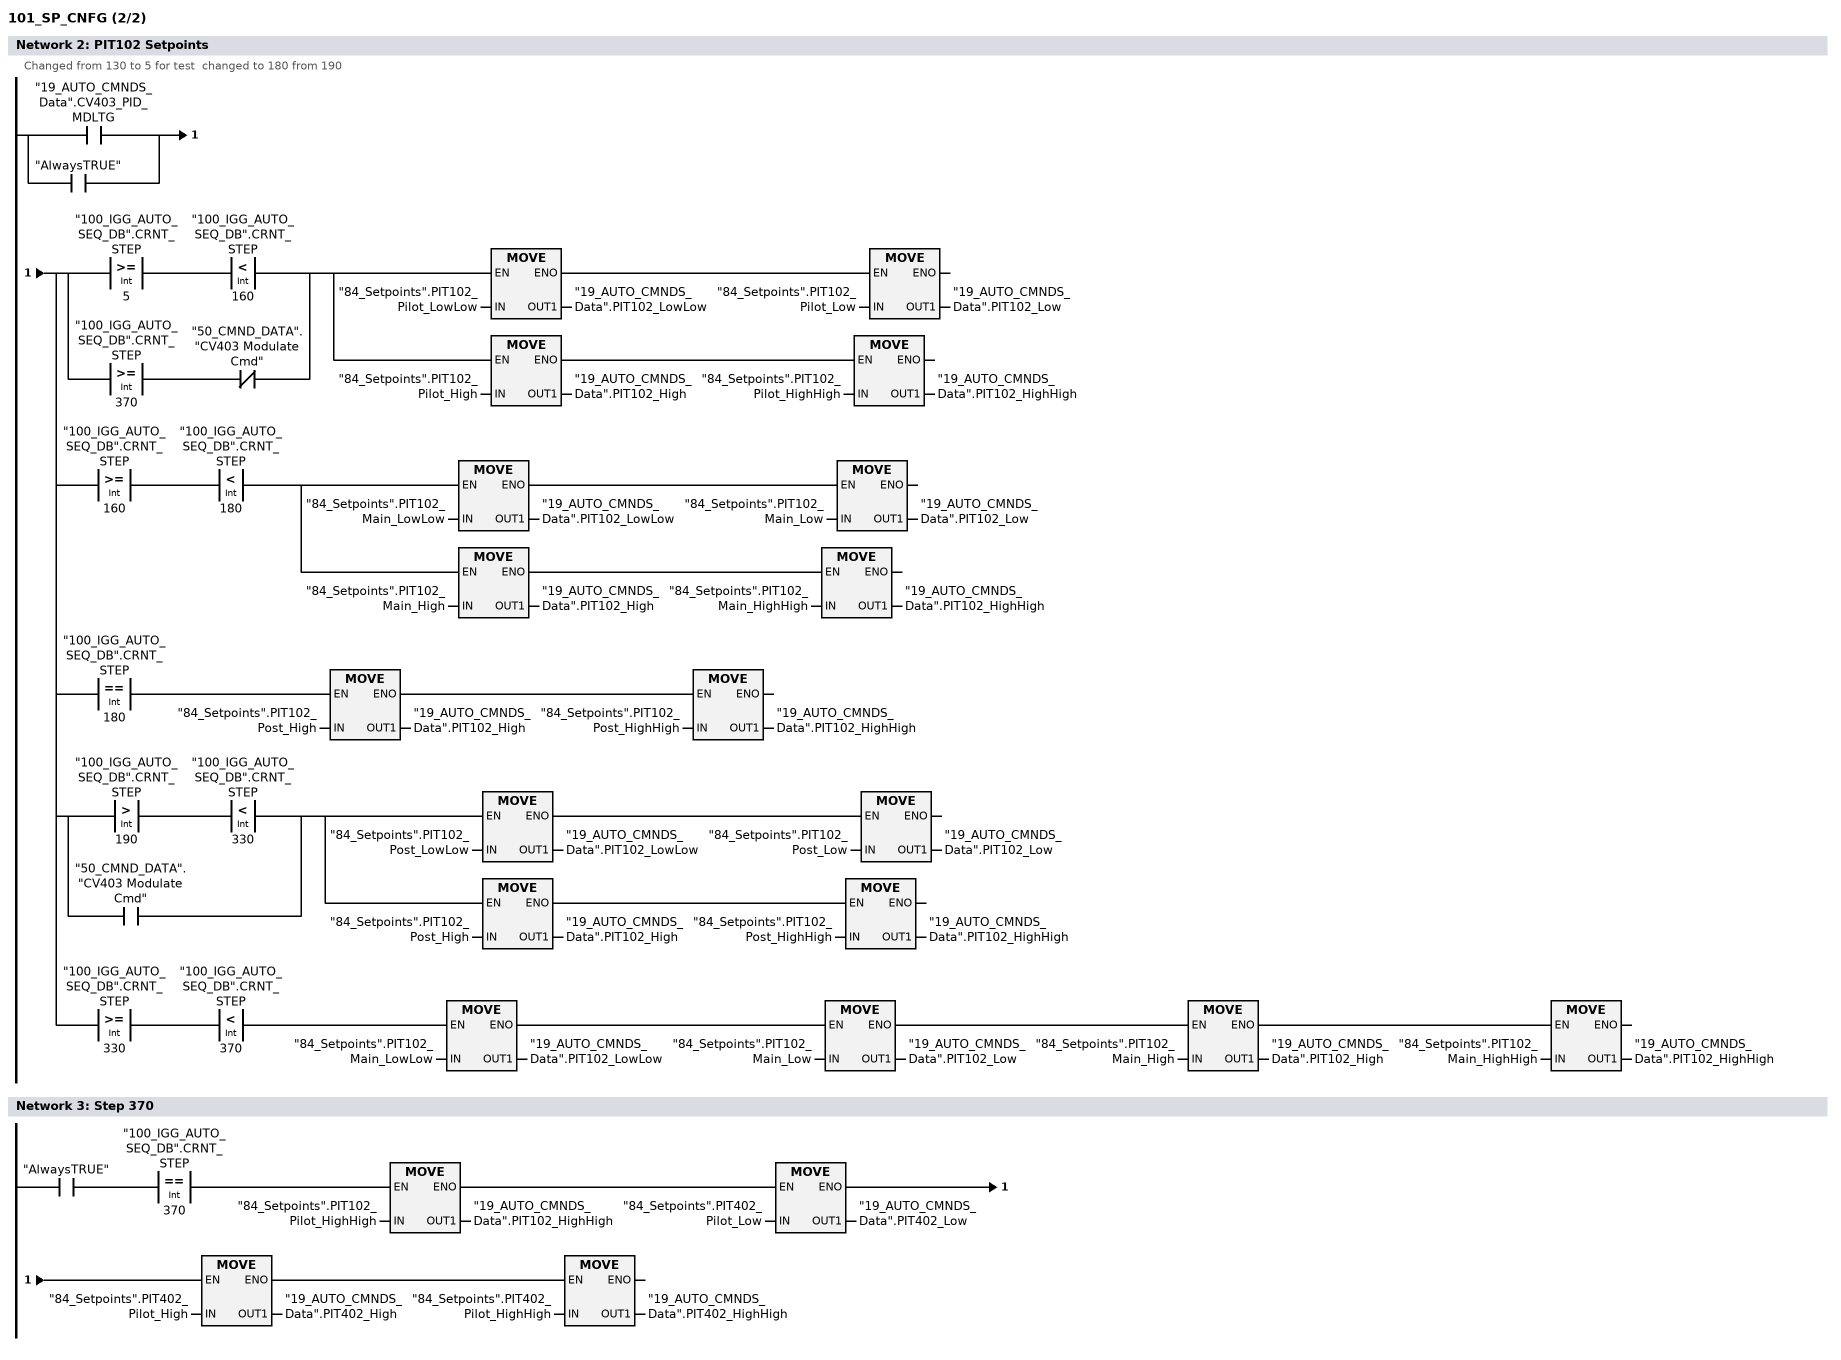
   RUNG wire#powerrail
      Contact( "19_AUTO_CMNDS_Data".CV403_PID_MDLTG )
      wire#w1
      { S7_Templates := "SrcType := Int" } GE_Contact(in1 := "100_IGG_AUTO_SEQ_DB".CRNT_STEP, in2 := 5)
      { S7_Templates := "SrcType := Int" } LT_Contact(in1 := "100_IGG_AUTO_SEQ_DB".CRNT_STEP, in2 := 160)
      wire#w2
      Move(in := "84_Setpoints".PIT102_Pilot_LowLow, out1 => "19_AUTO_CMNDS_Data".PIT102_LowLow)
      Move(in := "84_Setpoints".PIT102_Pilot_Low, out1 => "19_AUTO_CMNDS_Data".PIT102_Low)
   END_RUNG
   RUNG wire#powerrail
      Contact( "AlwaysTRUE" )
   END_RUNG wire#w1
   RUNG wire#w1
      { S7_Templates := "SrcType := Int" } GE_Contact(in1 := "100_IGG_AUTO_SEQ_DB".CRNT_STEP, in2 := 370)
      I_Contact( "50_CMND_DATA"."CV403 Modulate Cmd" )
   END_RUNG wire#w2
   RUNG wire#w2
      Move(in := "84_Setpoints".PIT102_Pilot_High, out1 => "19_AUTO_CMNDS_Data".PIT102_High)
      Move(in := "84_Setpoints".PIT102_Pilot_HighHigh, out1 => "19_AUTO_CMNDS_Data".PIT102_HighHigh)
   END_RUNG
   RUNG wire#w1
      { S7_Templates := "SrcType := Int" } GE_Contact(in1 := "100_IGG_AUTO_SEQ_DB".CRNT_STEP, in2 := 160)
      { S7_Templates := "SrcType := Int" } LT_Contact(in1 := "100_IGG_AUTO_SEQ_DB".CRNT_STEP, in2 := 180)
      wire#w3
      Move(in := "84_Setpoints".PIT102_Main_LowLow, out1 => "19_AUTO_CMNDS_Data".PIT102_LowLow)
      Move(in := "84_Setpoints".PIT102_Main_Low, out1 => "19_AUTO_CMNDS_Data".PIT102_Low)
   END_RUNG
   RUNG wire#w3
      Move(in := "84_Setpoints".PIT102_Main_High, out1 => "19_AUTO_CMNDS_Data".PIT102_High)
      Move(in := "84_Setpoints".PIT102_Main_HighHigh, out1 => "19_AUTO_CMNDS_Data".PIT102_HighHigh)
   END_RUNG
   RUNG wire#w1
      { S7_Templates := "SrcType := Int" } EQ_Contact(in1 := "100_IGG_AUTO_SEQ_DB".CRNT_STEP, in2 := 180)
      Move(in := "84_Setpoints".PIT102_Post_High, out1 => "19_AUTO_CMNDS_Data".PIT102_High)
      Move(in := "84_Setpoints".PIT102_Post_HighHigh, out1 => "19_AUTO_CMNDS_Data".PIT102_HighHigh)
   END_RUNG
   RUNG wire#w1
      { S7_Templates := "SrcType := Int" } GT_Contact(in1 := "100_IGG_AUTO_SEQ_DB".CRNT_STEP, in2 := 190)
      { S7_Templates := "SrcType := Int" } LT_Contact(in1 := "100_IGG_AUTO_SEQ_DB".CRNT_STEP, in2 := 330)
      wire#w4
      Move(in := "84_Setpoints".PIT102_Post_LowLow, out1 => "19_AUTO_CMNDS_Data".PIT102_LowLow)
      Move(in := "84_Setpoints".PIT102_Post_Low, out1 => "19_AUTO_CMNDS_Data".PIT102_Low)
   END_RUNG
   RUNG wire#w1
      Contact( "50_CMND_DATA"."CV403 Modulate Cmd" )
   END_RUNG wire#w4
   RUNG wire#w4
      Move(in := "84_Setpoints".PIT102_Post_High, out1 => "19_AUTO_CMNDS_Data".PIT102_High)
      Move(in := "84_Setpoints".PIT102_Post_HighHigh, out1 => "19_AUTO_CMNDS_Data".PIT102_HighHigh)
   END_RUNG
   RUNG wire#w1
      { S7_Templates := "SrcType := Int" } GE_Contact(in1 := "100_IGG_AUTO_SEQ_DB".CRNT_STEP, in2 := 330)
      { S7_Templates := "SrcType := Int" } LT_Contact(in1 := "100_IGG_AUTO_SEQ_DB".CRNT_STEP, in2 := 370)
      Move(in := "84_Setpoints".PIT102_Main_LowLow, out1 => "19_AUTO_CMNDS_Data".PIT102_LowLow)
      Move(in := "84_Setpoints".PIT102_Main_Low, out1 => "19_AUTO_CMNDS_Data".PIT102_Low)
      Move(in := "84_Setpoints".PIT102_Main_High, out1 => "19_AUTO_CMNDS_Data".PIT102_High)
      Move(in := "84_Setpoints".PIT102_Main_HighHigh, out1 => "19_AUTO_CMNDS_Data".PIT102_HighHigh)
   END_RUNG
   // the same network as SCL:
   #_w1 := "19_AUTO_CMNDS_Data".CV403_PID_MDLTG OR "AlwaysTRUE";
   IF #_w1 AND ((("100_IGG_AUTO_SEQ_DB".CRNT_STEP >= 5) AND ("100_IGG_AUTO_SEQ_DB".CRNT_STEP < 160)) OR (("100_IGG_AUTO_SEQ_DB".CRNT_STEP >= 370) AND NOT "50_CMND_DATA"."CV403 Modulate Cmd")) THEN
       "19_AUTO_CMNDS_Data".PIT102_LowLow := "84_Setpoints".PIT102_Pilot_LowLow;
       "19_AUTO_CMNDS_Data".PIT102_Low := "84_Setpoints".PIT102_Pilot_Low;
       "19_AUTO_CMNDS_Data".PIT102_High := "84_Setpoints".PIT102_Pilot_High;
       "19_AUTO_CMNDS_Data".PIT102_HighHigh := "84_Setpoints".PIT102_Pilot_HighHigh;
   END_IF;
   IF #_w1 AND ("100_IGG_AUTO_SEQ_DB".CRNT_STEP >= 160) AND ("100_IGG_AUTO_SEQ_DB".CRNT_STEP < 180) THEN
       "19_AUTO_CMNDS_Data".PIT102_LowLow := "84_Setpoints".PIT102_Main_LowLow;
       "19_AUTO_CMNDS_Data".PIT102_Low := "84_Setpoints".PIT102_Main_Low;
       "19_AUTO_CMNDS_Data".PIT102_High := "84_Setpoints".PIT102_Main_High;
       "19_AUTO_CMNDS_Data".PIT102_HighHigh := "84_Setpoints".PIT102_Main_HighHigh;
   END_IF;
   IF #_w1 AND ("100_IGG_AUTO_SEQ_DB".CRNT_STEP = 180) THEN
       "19_AUTO_CMNDS_Data".PIT102_High := "84_Setpoints".PIT102_Post_High;
       "19_AUTO_CMNDS_Data".PIT102_HighHigh := "84_Setpoints".PIT102_Post_HighHigh;
   END_IF;
   IF #_w1 AND ((("100_IGG_AUTO_SEQ_DB".CRNT_STEP > 190) AND ("100_IGG_AUTO_SEQ_DB".CRNT_STEP < 330)) OR "50_CMND_DATA"."CV403 Modulate Cmd") THEN
       "19_AUTO_CMNDS_Data".PIT102_LowLow := "84_Setpoints".PIT102_Post_LowLow;
       "19_AUTO_CMNDS_Data".PIT102_Low := "84_Setpoints".PIT102_Post_Low;
       "19_AUTO_CMNDS_Data".PIT102_High := "84_Setpoints".PIT102_Post_High;
       "19_AUTO_CMNDS_Data".PIT102_HighHigh := "84_Setpoints".PIT102_Post_HighHigh;
   END_IF;
   IF #_w1 AND ("100_IGG_AUTO_SEQ_DB".CRNT_STEP >= 330) AND ("100_IGG_AUTO_SEQ_DB".CRNT_STEP < 370) THEN
       "19_AUTO_CMNDS_Data".PIT102_LowLow := "84_Setpoints".PIT102_Main_LowLow;
       "19_AUTO_CMNDS_Data".PIT102_Low := "84_Setpoints".PIT102_Main_Low;
       "19_AUTO_CMNDS_Data".PIT102_High := "84_Setpoints".PIT102_Main_High;
       "19_AUTO_CMNDS_Data".PIT102_HighHigh := "84_Setpoints".PIT102_Main_HighHigh;
   END_IF;
END_REGION

REGION Network 3: Step 370
   RUNG wire#powerrail
      Contact( "AlwaysTRUE" )
      { S7_Templates := "SrcType := Int" } EQ_Contact(in1 := "100_IGG_AUTO_SEQ_DB".CRNT_STEP, in2 := 370)
      Move(in := "84_Setpoints".PIT102_Pilot_HighHigh, out1 => "19_AUTO_CMNDS_Data".PIT102_HighHigh)
      Move(in := "84_Setpoints".PIT402_Pilot_Low, out1 => "19_AUTO_CMNDS_Data".PIT402_Low)
      Move(in := "84_Setpoints".PIT402_Pilot_High, out1 => "19_AUTO_CMNDS_Data".PIT402_High)
      Move(in := "84_Setpoints".PIT402_Pilot_HighHigh, out1 => "19_AUTO_CMNDS_Data".PIT402_HighHigh)
   END_RUNG
   // the same network as SCL:
   IF "AlwaysTRUE" AND ("100_IGG_AUTO_SEQ_DB".CRNT_STEP = 370) THEN
       "19_AUTO_CMNDS_Data".PIT102_HighHigh := "84_Setpoints".PIT102_Pilot_HighHigh;
       "19_AUTO_CMNDS_Data".PIT402_Low := "84_Setpoints".PIT402_Pilot_Low;
       "19_AUTO_CMNDS_Data".PIT402_High := "84_Setpoints".PIT402_Pilot_High;
       "19_AUTO_CMNDS_Data".PIT402_HighHigh := "84_Setpoints".PIT402_Pilot_HighHigh;
   END_IF;
END_REGION
END_FUNCTION

// folder: 120 - 139 FAT Functions

FUNCTION "120_FAT_FCS" : Void   // FC120, LAD
TITLE = FAT Functions
{ S7_Optimized_Access := 'TRUE' }
AUTHOR : JRS
VERSION : 0.1
// For specific functions related to the factory test equipment & setup
   VAR_TEMP   // added for the SCL form of the ladder/FBD networks
      _w1 : Bool;
   END_VAR
BEGIN

REGION Network 1: Into FAT Mode
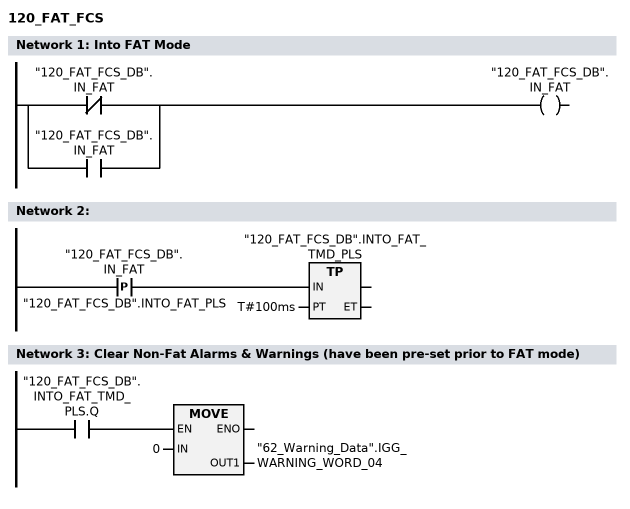
   RUNG wire#powerrail
      I_Contact( "120_FAT_FCS_DB".IN_FAT )
      wire#w1
      Coil( "120_FAT_FCS_DB".IN_FAT )
   END_RUNG
   RUNG wire#powerrail
      Contact( "120_FAT_FCS_DB".IN_FAT )
   END_RUNG wire#w1
   // the same network as SCL:
   "120_FAT_FCS_DB".IN_FAT := NOT "120_FAT_FCS_DB".IN_FAT OR "120_FAT_FCS_DB".IN_FAT;
END_REGION

REGION Network 2
   #_w1 := "120_FAT_FCS_DB".IN_FAT AND NOT "120_FAT_FCS_DB".INTO_FAT_PLS;   // rising edge of "120_FAT_FCS_DB".IN_FAT
   "120_FAT_FCS_DB".INTO_FAT_PLS := "120_FAT_FCS_DB".IN_FAT;
   "120_FAT_FCS_DB".INTO_FAT_TMD_PLS.TP(IN := #_w1, PT := T#100ms);
END_REGION

REGION Network 3: Clear Non-Fat Alarms & Warnings (have been pre-set prior to FAT mode)
   RUNG wire#powerrail
      Contact( "120_FAT_FCS_DB".INTO_FAT_TMD_PLS.Q )
      Move(in := 0, out1 => "62_Warning_Data".IGG_WARNING_WORD_04)
   END_RUNG
   // the same network as SCL:
   IF "120_FAT_FCS_DB".INTO_FAT_TMD_PLS.Q THEN "62_Warning_Data".IGG_WARNING_WORD_04 := 0; END_IF;
END_REGION
END_FUNCTION

// folder: 300 - 499 Counters and Timer DBs

FUNCTION "300_AUT_SUQ_TIMERS" : Void   // FC300, LAD
TITLE = Automatic Sequence Timers
{ S7_Optimized_Access := 'TRUE' }
AUTHOR : JRS
VERSION : 0.1
// For specific sequence timers not covered by step FB timers
BEGIN

REGION Network 1: Pre BC Start Command Delay
   // Get time value from HMI data
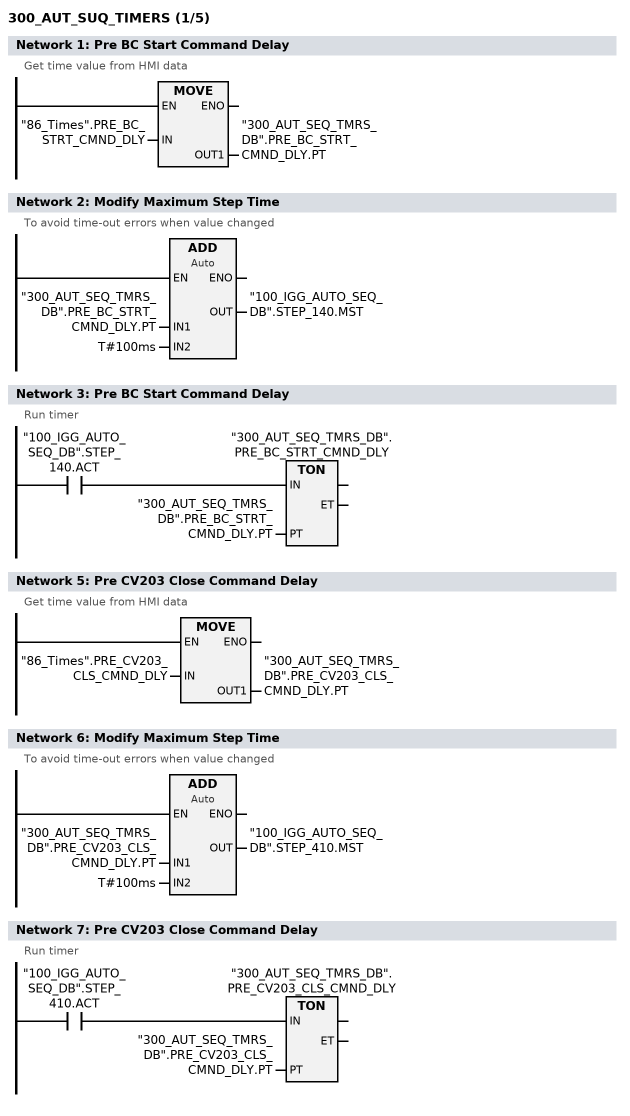
   RUNG wire#powerrail
      Move(in := "86_Times".PRE_BC_STRT_CMND_DLY, out1 => "300_AUT_SEQ_TMRS_DB".PRE_BC_STRT_CMND_DLY.PT)
   END_RUNG
   // the same network as SCL:
   "300_AUT_SEQ_TMRS_DB".PRE_BC_STRT_CMND_DLY.PT := "86_Times".PRE_BC_STRT_CMND_DLY;
END_REGION

REGION Network 2: Modify Maximum Step Time
   // To avoid time-out errors when value changed
   RUNG wire#powerrail
      Add(in1 := "300_AUT_SEQ_TMRS_DB".PRE_BC_STRT_CMND_DLY.PT, in2 := T#100ms, out => "100_IGG_AUTO_SEQ_DB".STEP_140.MST)
   END_RUNG
   // the same network as SCL:
   "100_IGG_AUTO_SEQ_DB".STEP_140.MST := "300_AUT_SEQ_TMRS_DB".PRE_BC_STRT_CMND_DLY.PT + T#100ms;
END_REGION

REGION Network 3: Pre BC Start Command Delay
   // Run timer
   "300_AUT_SEQ_TMRS_DB".PRE_BC_STRT_CMND_DLY.TON(IN := "100_IGG_AUTO_SEQ_DB".STEP_140.ACT,
                           PT := "300_AUT_SEQ_TMRS_DB".PRE_BC_STRT_CMND_DLY.PT);
END_REGION

REGION Network 5: Pre CV203 Close Command Delay
   // Get time value from HMI data
   RUNG wire#powerrail
      Move(in := "86_Times".PRE_CV203_CLS_CMND_DLY, out1 => "300_AUT_SEQ_TMRS_DB".PRE_CV203_CLS_CMND_DLY.PT)
   END_RUNG
   // the same network as SCL:
   "300_AUT_SEQ_TMRS_DB".PRE_CV203_CLS_CMND_DLY.PT := "86_Times".PRE_CV203_CLS_CMND_DLY;
END_REGION

REGION Network 6: Modify Maximum Step Time
   // To avoid time-out errors when value changed
   RUNG wire#powerrail
      Add(in1 := "300_AUT_SEQ_TMRS_DB".PRE_CV203_CLS_CMND_DLY.PT, in2 := T#100ms, out => "100_IGG_AUTO_SEQ_DB".STEP_410.MST)
   END_RUNG
   // the same network as SCL:
   "100_IGG_AUTO_SEQ_DB".STEP_410.MST := "300_AUT_SEQ_TMRS_DB".PRE_CV203_CLS_CMND_DLY.PT + T#100ms;
END_REGION

REGION Network 7: Pre CV203 Close Command Delay
   // Run timer
   "300_AUT_SEQ_TMRS_DB".PRE_CV203_CLS_CMND_DLY.TON(IN := "100_IGG_AUTO_SEQ_DB".STEP_410.ACT,
                           PT := "300_AUT_SEQ_TMRS_DB".PRE_CV203_CLS_CMND_DLY.PT);
END_REGION

REGION Network 9: Post P301 Stop Delay
   // Get time value from HMI data
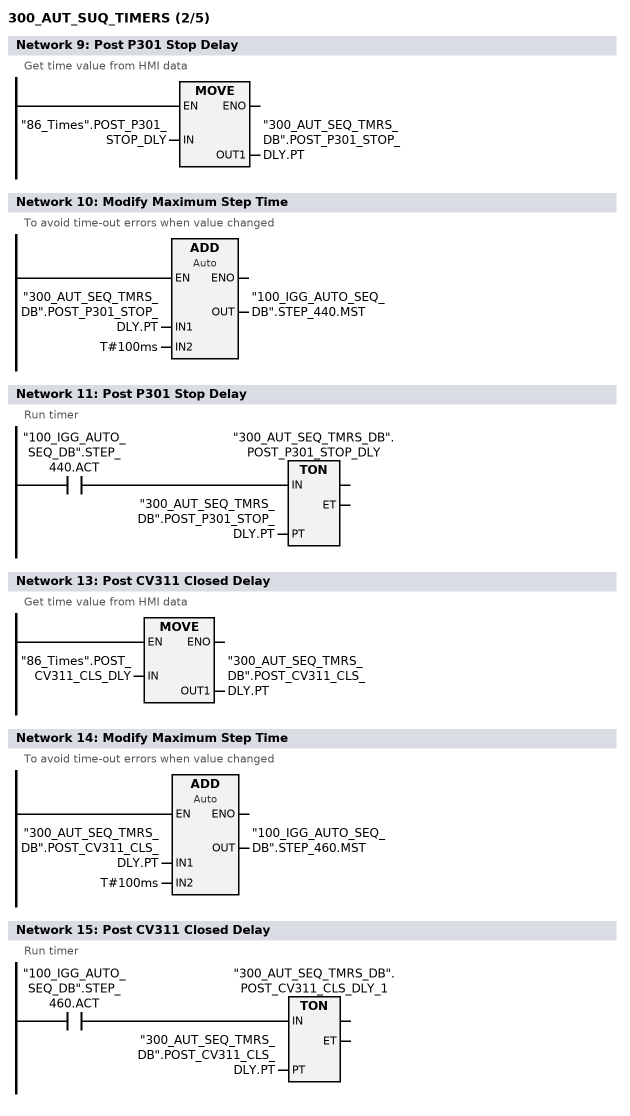
   RUNG wire#powerrail
      Move(in := "86_Times".POST_P301_STOP_DLY, out1 => "300_AUT_SEQ_TMRS_DB".POST_P301_STOP_DLY.PT)
   END_RUNG
   // the same network as SCL:
   "300_AUT_SEQ_TMRS_DB".POST_P301_STOP_DLY.PT := "86_Times".POST_P301_STOP_DLY;
END_REGION

REGION Network 10: Modify Maximum Step Time
   // To avoid time-out errors when value changed
   RUNG wire#powerrail
      Add(in1 := "300_AUT_SEQ_TMRS_DB".POST_P301_STOP_DLY.PT, in2 := T#100ms, out => "100_IGG_AUTO_SEQ_DB".STEP_440.MST)
   END_RUNG
   // the same network as SCL:
   "100_IGG_AUTO_SEQ_DB".STEP_440.MST := "300_AUT_SEQ_TMRS_DB".POST_P301_STOP_DLY.PT + T#100ms;
END_REGION

REGION Network 11: Post P301 Stop Delay
   // Run timer
   "300_AUT_SEQ_TMRS_DB".POST_P301_STOP_DLY.TON(IN := "100_IGG_AUTO_SEQ_DB".STEP_440.ACT,
                           PT := "300_AUT_SEQ_TMRS_DB".POST_P301_STOP_DLY.PT);
END_REGION

REGION Network 13: Post CV311 Closed Delay
   // Get time value from HMI data
   RUNG wire#powerrail
      Move(in := "86_Times".POST_CV311_CLS_DLY, out1 => "300_AUT_SEQ_TMRS_DB".POST_CV311_CLS_DLY.PT)
   END_RUNG
   // the same network as SCL:
   "300_AUT_SEQ_TMRS_DB".POST_CV311_CLS_DLY.PT := "86_Times".POST_CV311_CLS_DLY;
END_REGION

REGION Network 14: Modify Maximum Step Time
   // To avoid time-out errors when value changed
   RUNG wire#powerrail
      Add(in1 := "300_AUT_SEQ_TMRS_DB".POST_CV311_CLS_DLY.PT, in2 := T#100ms, out => "100_IGG_AUTO_SEQ_DB".STEP_460.MST)
   END_RUNG
   // the same network as SCL:
   "100_IGG_AUTO_SEQ_DB".STEP_460.MST := "300_AUT_SEQ_TMRS_DB".POST_CV311_CLS_DLY.PT + T#100ms;
END_REGION

REGION Network 15: Post CV311 Closed Delay
   // Run timer
   "300_AUT_SEQ_TMRS_DB".POST_CV311_CLS_DLY_1.TON(IN := "100_IGG_AUTO_SEQ_DB".STEP_460.ACT,
                           PT := "300_AUT_SEQ_TMRS_DB".POST_CV311_CLS_DLY.PT);
END_REGION

REGION Network 17: Post CV321 Opened Delay
   // Get time value from HMI data
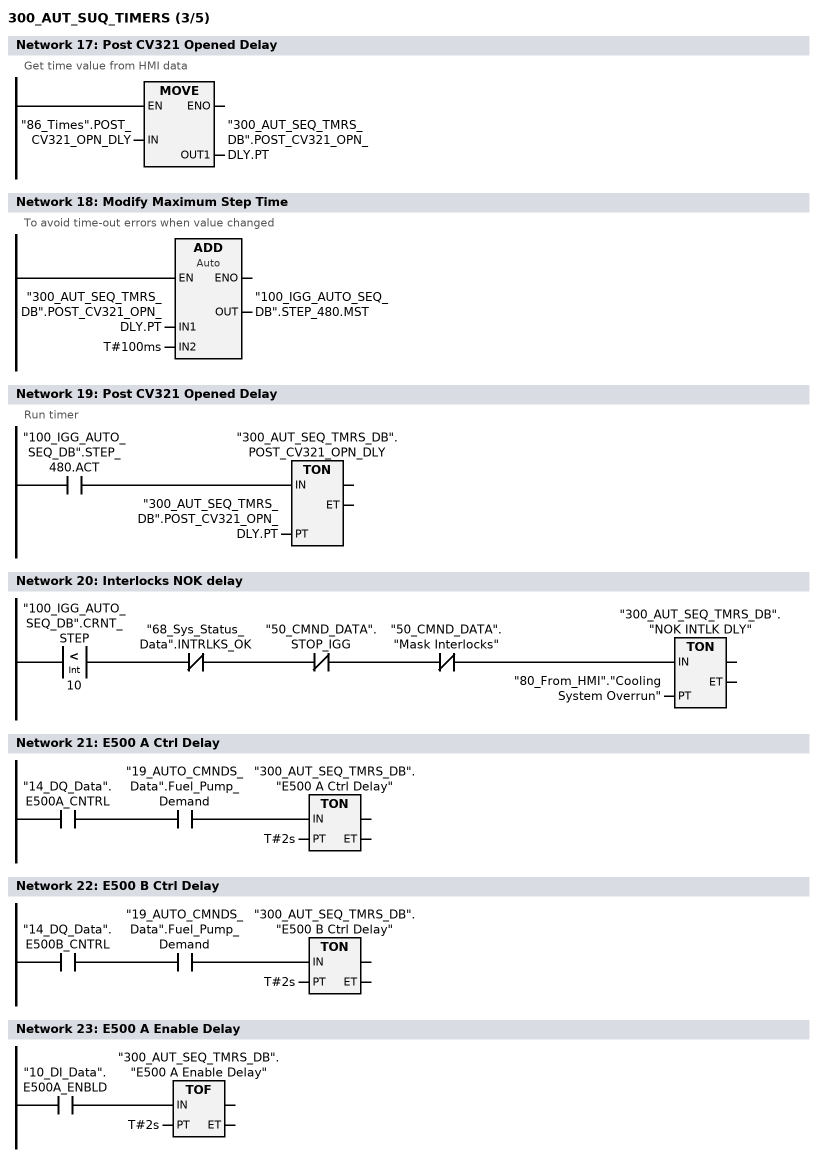
   RUNG wire#powerrail
      Move(in := "86_Times".POST_CV321_OPN_DLY, out1 => "300_AUT_SEQ_TMRS_DB".POST_CV321_OPN_DLY.PT)
   END_RUNG
   // the same network as SCL:
   "300_AUT_SEQ_TMRS_DB".POST_CV321_OPN_DLY.PT := "86_Times".POST_CV321_OPN_DLY;
END_REGION

REGION Network 18: Modify Maximum Step Time
   // To avoid time-out errors when value changed
   RUNG wire#powerrail
      Add(in1 := "300_AUT_SEQ_TMRS_DB".POST_CV321_OPN_DLY.PT, in2 := T#100ms, out => "100_IGG_AUTO_SEQ_DB".STEP_480.MST)
   END_RUNG
   // the same network as SCL:
   "100_IGG_AUTO_SEQ_DB".STEP_480.MST := "300_AUT_SEQ_TMRS_DB".POST_CV321_OPN_DLY.PT + T#100ms;
END_REGION

REGION Network 19: Post CV321 Opened Delay
   // Run timer
   "300_AUT_SEQ_TMRS_DB".POST_CV321_OPN_DLY.TON(IN := "100_IGG_AUTO_SEQ_DB".STEP_480.ACT,
                           PT := "300_AUT_SEQ_TMRS_DB".POST_CV321_OPN_DLY.PT);
END_REGION

REGION Network 20: Interlocks NOK delay
   "300_AUT_SEQ_TMRS_DB"."NOK INTLK DLY".TON(IN := ("100_IGG_AUTO_SEQ_DB".CRNT_STEP < 10) AND NOT "68_Sys_Status_Data".INTRLKS_OK AND NOT "50_CMND_DATA".STOP_IGG AND NOT "50_CMND_DATA"."Mask Interlocks",
                           PT := "80_From_HMI"."Cooling System Overrun");
END_REGION

REGION Network 21: E500 A Ctrl Delay
   "300_AUT_SEQ_TMRS_DB"."E500 A Ctrl Delay".TON(IN := "14_DQ_Data".E500A_CNTRL AND "19_AUTO_CMNDS_Data".Fuel_Pump_Demand,
                           PT := T#2s);
END_REGION

REGION Network 22: E500 B Ctrl Delay
   "300_AUT_SEQ_TMRS_DB"."E500 B Ctrl Delay".TON(IN := "14_DQ_Data".E500B_CNTRL AND "19_AUTO_CMNDS_Data".Fuel_Pump_Demand,
                           PT := T#2s);
END_REGION

REGION Network 23: E500 A Enable Delay
   "300_AUT_SEQ_TMRS_DB"."E500 A Enable Delay".TOF(IN := "10_DI_Data".E500A_ENBLD, PT := T#2s);
END_REGION

REGION Network 24: E500 B Enable Delay
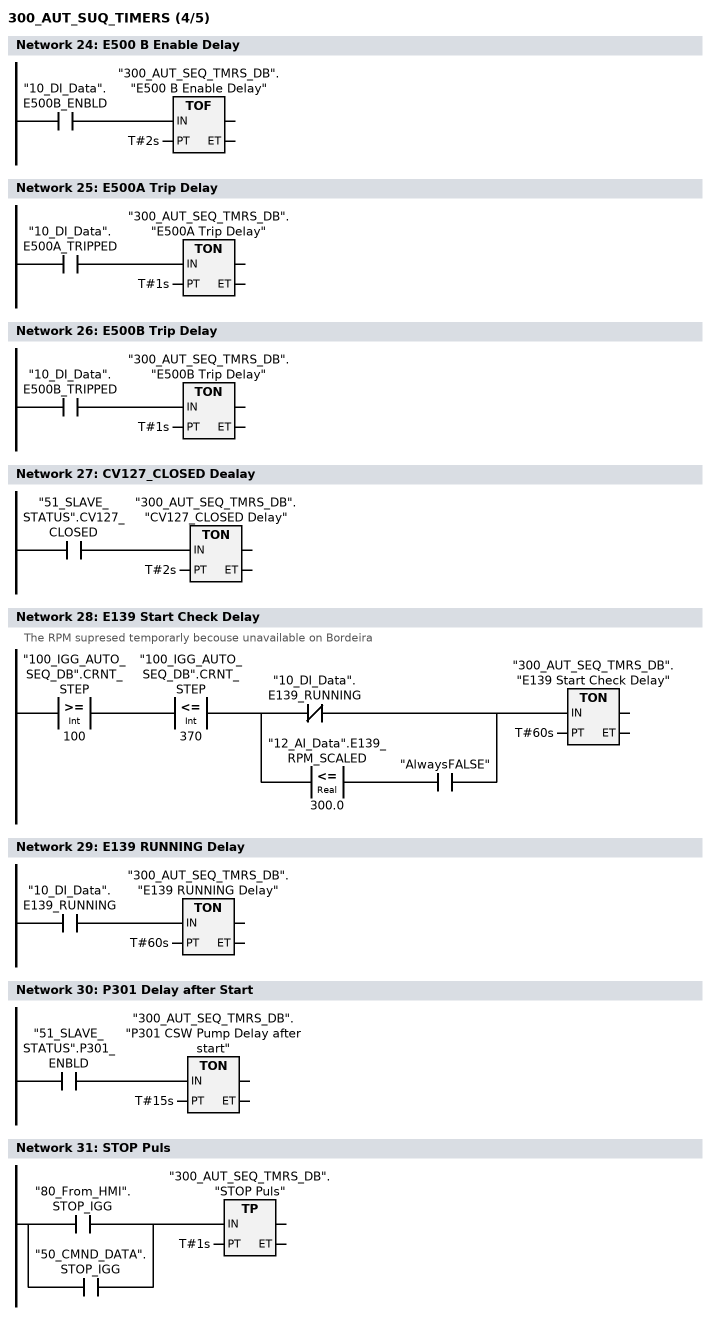
   "300_AUT_SEQ_TMRS_DB"."E500 B Enable Delay".TOF(IN := "10_DI_Data".E500B_ENBLD, PT := T#2s);
END_REGION

REGION Network 25: E500A Trip Delay
   "300_AUT_SEQ_TMRS_DB"."E500A Trip Delay".TON(IN := "10_DI_Data".E500A_TRIPPED, PT := T#1s);
END_REGION

REGION Network 26: E500B Trip Delay
   "300_AUT_SEQ_TMRS_DB"."E500B Trip Delay".TON(IN := "10_DI_Data".E500B_TRIPPED, PT := T#1s);
END_REGION

REGION Network 27: CV127_CLOSED Dealay
   "300_AUT_SEQ_TMRS_DB"."CV127_CLOSED Delay".TON(IN := "51_SLAVE_STATUS".CV127_CLOSED, PT := T#2s);
END_REGION

REGION Network 28: E139 Start Check Delay
   // The RPM supresed temporarly becouse unavailable on Bordeira
   "300_AUT_SEQ_TMRS_DB"."E139 Start Check Delay".TON(IN := ("100_IGG_AUTO_SEQ_DB".CRNT_STEP >= 100) AND ("100_IGG_AUTO_SEQ_DB".CRNT_STEP <= 370) AND (NOT "10_DI_Data".E139_RUNNING OR (("12_AI_Data".E139_RPM_SCALED <= 300.0) AND "AlwaysFALSE")),
                           PT := T#60s);
END_REGION

REGION Network 29: E139 RUNNING Delay
   "300_AUT_SEQ_TMRS_DB"."E139 RUNNING Delay".TON(IN := "10_DI_Data".E139_RUNNING, PT := T#60s);
END_REGION

REGION Network 30: P301 Delay after Start
   "300_AUT_SEQ_TMRS_DB"."P301 CSW Pump Delay after start".TON(IN := "51_SLAVE_STATUS".P301_ENBLD, PT := T#15s);
END_REGION

REGION Network 31: STOP Puls
   "300_AUT_SEQ_TMRS_DB"."STOP Puls".TP(IN := "80_From_HMI".STOP_IGG OR "50_CMND_DATA".STOP_IGG, PT := T#1s);
END_REGION

REGION Network 32: E-Stop Loop
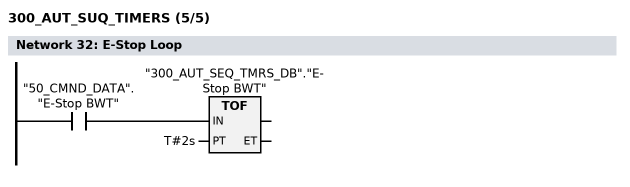
   "300_AUT_SEQ_TMRS_DB"."E-Stop BWT".TOF(IN := "50_CMND_DATA"."E-Stop BWT", PT := T#2s);
END_REGION
END_FUNCTION

// folder: 50 - 59 Communication

FUNCTION "51_GET_SLAVE_DATA" : Void   // FC51, LAD
TITLE = Get Slave Status Data
{ S7_Optimized_Access := 'TRUE' }
AUTHOR : JRS
VERSION : 0.1
// Code for getting status data from the slave PLC
BEGIN

REGION Network 1: Get Slave Status Data
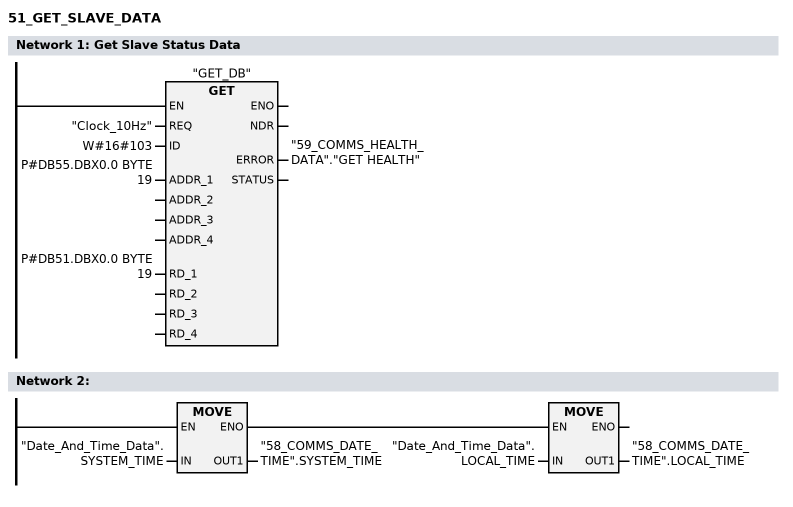
   "GET_DB"(REQ := "Clock_10Hz",   // GET
            ID := W#16#103,
            ADDR_1 := P#DB55.DBX0.0 BYTE 19,
            RD_1 := P#DB51.DBX0.0 BYTE 19,
            ERROR => "59_COMMS_HEALTH_DATA"."GET HEALTH");
END_REGION

REGION Network 2
   RUNG wire#powerrail
      Move(in := "Date_And_Time_Data".SYSTEM_TIME, out1 => "58_COMMS_DATE_TIME".SYSTEM_TIME)
      Move(in := "Date_And_Time_Data".LOCAL_TIME, out1 => "58_COMMS_DATE_TIME".LOCAL_TIME)
   END_RUNG
   // the same network as SCL:
   "58_COMMS_DATE_TIME".SYSTEM_TIME := "Date_And_Time_Data".SYSTEM_TIME;
   "58_COMMS_DATE_TIME".LOCAL_TIME := "Date_And_Time_Data".LOCAL_TIME;
END_REGION
END_FUNCTION

FUNCTION "56_PUT_SLAVE_DATA" : Void   // FC56, LAD
TITLE = Put Slave Comands Data
{ S7_Optimized_Access := 'TRUE' }
AUTHOR : JRS
VERSION : 0.1
// Code for sending commands to the slave PLC
   VAR_TEMP
      RACK_2_done : Bool;
      RACK_2_error : Bool;
      RACK_2_status : Word;
      RACK_3_done : Bool;
      RACK_3_error : Bool;
      RACK_3_status : Word;
   END_VAR
BEGIN

REGION Network 1: PUT Slave Commands
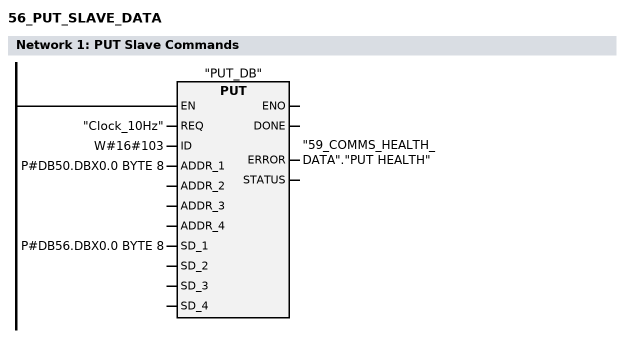
   "PUT_DB"(REQ := "Clock_10Hz",   // PUT
            ID := W#16#103,
            ADDR_1 := P#DB50.DBX0.0 BYTE 8,
            SD_1 := P#DB56.DBX0.0 BYTE 8,
            ERROR => "59_COMMS_HEALTH_DATA"."PUT HEALTH");
END_REGION
END_FUNCTION

FUNCTION "59_COMMS_HEALTH" : Void   // FC59, LAD
TITLE = Communications Heart Beats
{ S7_Optimized_Access := 'TRUE' }
AUTHOR : JRS
VERSION : 0.1
// Code for communications health determination
   VAR_TEMP   // added for the SCL form of the ladder/FBD networks
      _w1 : Bool;
      _w2 : Bool;
   END_VAR
BEGIN

REGION Network 1: Local Heart Beat
   // Flip flop for status to other PLC's
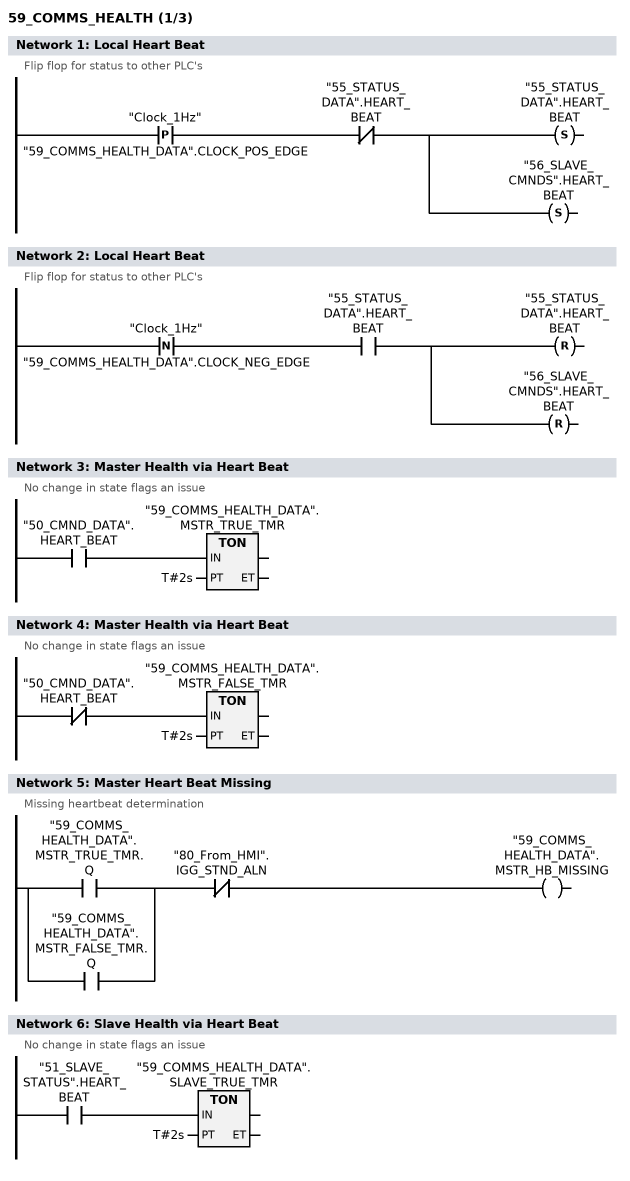
   RUNG wire#powerrail
      P_Contact(operand := "Clock_1Hz", bit := "59_COMMS_HEALTH_DATA".CLOCK_POS_EDGE)
      I_Contact( "55_STATUS_DATA".HEART_BEAT )
      wire#w1
      S_Coil( "55_STATUS_DATA".HEART_BEAT )
   END_RUNG
   RUNG wire#w1
      S_Coil( "56_SLAVE_CMNDS".HEART_BEAT )
   END_RUNG
   // the same network as SCL:
   #_w1 := "Clock_1Hz" AND NOT "59_COMMS_HEALTH_DATA".CLOCK_POS_EDGE;   // rising edge of "Clock_1Hz"
   "59_COMMS_HEALTH_DATA".CLOCK_POS_EDGE := "Clock_1Hz";
   #_w2 := #_w1 AND NOT "55_STATUS_DATA".HEART_BEAT;
   IF #_w2 THEN
       "55_STATUS_DATA".HEART_BEAT := TRUE;
       "56_SLAVE_CMNDS".HEART_BEAT := TRUE;
   END_IF;
END_REGION

REGION Network 2: Local Heart Beat
   // Flip flop for status to other PLC's
   RUNG wire#powerrail
      N_Contact(operand := "Clock_1Hz", bit := "59_COMMS_HEALTH_DATA".CLOCK_NEG_EDGE)
      Contact( "55_STATUS_DATA".HEART_BEAT )
      wire#w1
      R_Coil( "55_STATUS_DATA".HEART_BEAT )
   END_RUNG
   RUNG wire#w1
      R_Coil( "56_SLAVE_CMNDS".HEART_BEAT )
   END_RUNG
   // the same network as SCL:
   #_w1 := NOT "Clock_1Hz" AND "59_COMMS_HEALTH_DATA".CLOCK_NEG_EDGE;   // falling edge of "Clock_1Hz"
   "59_COMMS_HEALTH_DATA".CLOCK_NEG_EDGE := "Clock_1Hz";
   #_w2 := #_w1 AND "55_STATUS_DATA".HEART_BEAT;
   IF #_w2 THEN
       "55_STATUS_DATA".HEART_BEAT := FALSE;
       "56_SLAVE_CMNDS".HEART_BEAT := FALSE;
   END_IF;
END_REGION

REGION Network 3: Master Health via Heart Beat
   // No change in state flags an issue
   "59_COMMS_HEALTH_DATA".MSTR_TRUE_TMR.TON(IN := "50_CMND_DATA".HEART_BEAT, PT := T#2s);
END_REGION

REGION Network 4: Master Health via Heart Beat
   // No change in state flags an issue
   "59_COMMS_HEALTH_DATA".MSTR_FALSE_TMR.TON(IN := NOT "50_CMND_DATA".HEART_BEAT, PT := T#2s);
END_REGION

REGION Network 5: Master Heart Beat Missing
   // Missing heartbeat determination
   RUNG wire#powerrail
      Contact( "59_COMMS_HEALTH_DATA".MSTR_TRUE_TMR.Q )
      wire#w1
      I_Contact( "80_From_HMI".IGG_STND_ALN )
      Coil( "59_COMMS_HEALTH_DATA".MSTR_HB_MISSING )
   END_RUNG
   RUNG wire#powerrail
      Contact( "59_COMMS_HEALTH_DATA".MSTR_FALSE_TMR.Q )
   END_RUNG wire#w1
   // the same network as SCL:
   "59_COMMS_HEALTH_DATA".MSTR_HB_MISSING := ("59_COMMS_HEALTH_DATA".MSTR_TRUE_TMR.Q OR "59_COMMS_HEALTH_DATA".MSTR_FALSE_TMR.Q) AND NOT "80_From_HMI".IGG_STND_ALN;
END_REGION

REGION Network 6: Slave Health via Heart Beat
   // No change in state flags an issue
   "59_COMMS_HEALTH_DATA".SLAVE_TRUE_TMR.TON(IN := "51_SLAVE_STATUS".HEART_BEAT, PT := T#2s);
END_REGION

REGION Network 7: Slave Health via Heart Beat
   // No change in state flags an issue
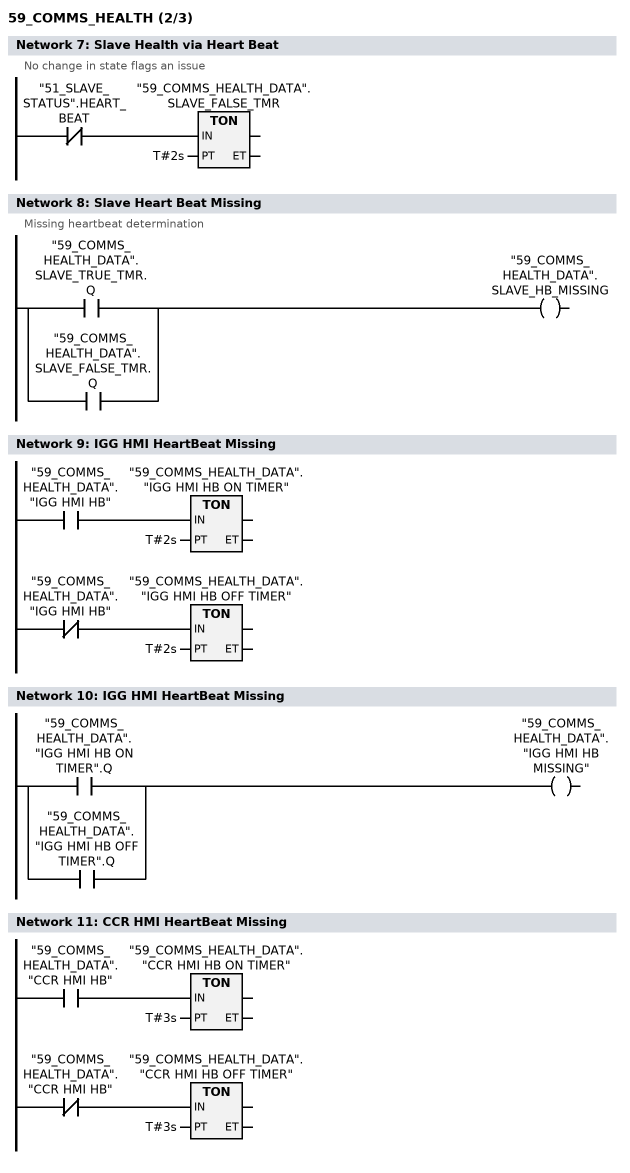
   "59_COMMS_HEALTH_DATA".SLAVE_FALSE_TMR.TON(IN := NOT "51_SLAVE_STATUS".HEART_BEAT, PT := T#2s);
END_REGION

REGION Network 8: Slave Heart Beat Missing
   // Missing heartbeat determination
   RUNG wire#powerrail
      Contact( "59_COMMS_HEALTH_DATA".SLAVE_TRUE_TMR.Q )
      wire#w1
      Coil( "59_COMMS_HEALTH_DATA".SLAVE_HB_MISSING )
   END_RUNG
   RUNG wire#powerrail
      Contact( "59_COMMS_HEALTH_DATA".SLAVE_FALSE_TMR.Q )
   END_RUNG wire#w1
   // the same network as SCL:
   "59_COMMS_HEALTH_DATA".SLAVE_HB_MISSING := "59_COMMS_HEALTH_DATA".SLAVE_TRUE_TMR.Q OR "59_COMMS_HEALTH_DATA".SLAVE_FALSE_TMR.Q;
END_REGION

REGION Network 9: IGG HMI HeartBeat Missing
   "59_COMMS_HEALTH_DATA"."IGG HMI HB ON TIMER".TON(IN := "59_COMMS_HEALTH_DATA"."IGG HMI HB", PT := T#2s);
   "59_COMMS_HEALTH_DATA"."IGG HMI HB OFF TIMER".TON(IN := NOT "59_COMMS_HEALTH_DATA"."IGG HMI HB", PT := T#2s);
END_REGION

REGION Network 10: IGG HMI HeartBeat Missing
   RUNG wire#powerrail
      Contact( "59_COMMS_HEALTH_DATA"."IGG HMI HB ON TIMER".Q )
      wire#w1
      Coil( "59_COMMS_HEALTH_DATA"."IGG HMI HB MISSING" )
   END_RUNG
   RUNG wire#powerrail
      Contact( "59_COMMS_HEALTH_DATA"."IGG HMI HB OFF TIMER".Q )
   END_RUNG wire#w1
   // the same network as SCL:
   "59_COMMS_HEALTH_DATA"."IGG HMI HB MISSING" := "59_COMMS_HEALTH_DATA"."IGG HMI HB ON TIMER".Q OR "59_COMMS_HEALTH_DATA"."IGG HMI HB OFF TIMER".Q;
END_REGION

REGION Network 11: CCR HMI HeartBeat Missing
   "59_COMMS_HEALTH_DATA"."CCR HMI HB ON TIMER".TON(IN := "59_COMMS_HEALTH_DATA"."CCR HMI HB", PT := T#3s);
   "59_COMMS_HEALTH_DATA"."CCR HMI HB OFF TIMER".TON(IN := NOT "59_COMMS_HEALTH_DATA"."CCR HMI HB", PT := T#3s);
END_REGION

REGION Network 12: CCR HMI HeartBeat Missing
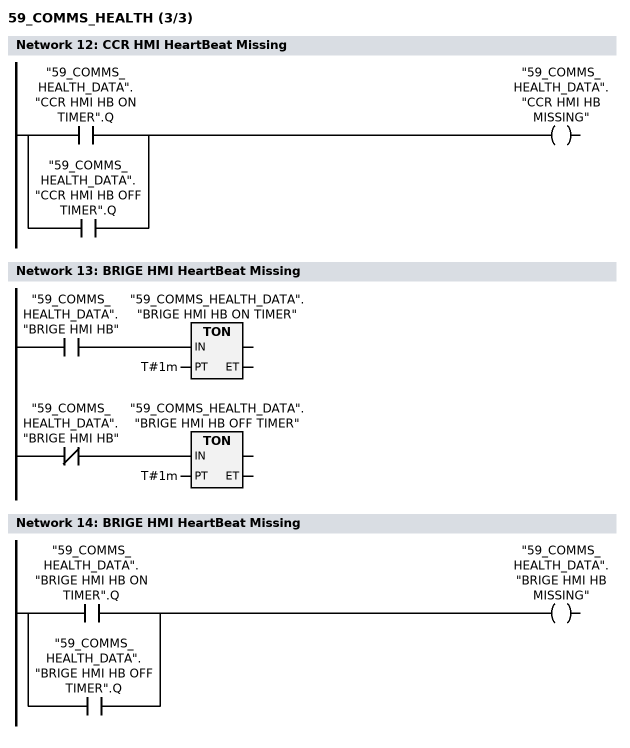
   RUNG wire#powerrail
      Contact( "59_COMMS_HEALTH_DATA"."CCR HMI HB ON TIMER".Q )
      wire#w1
      Coil( "59_COMMS_HEALTH_DATA"."CCR HMI HB MISSING" )
   END_RUNG
   RUNG wire#powerrail
      Contact( "59_COMMS_HEALTH_DATA"."CCR HMI HB OFF TIMER".Q )
   END_RUNG wire#w1
   // the same network as SCL:
   "59_COMMS_HEALTH_DATA"."CCR HMI HB MISSING" := "59_COMMS_HEALTH_DATA"."CCR HMI HB ON TIMER".Q OR "59_COMMS_HEALTH_DATA"."CCR HMI HB OFF TIMER".Q;
END_REGION

REGION Network 13: BRIGE HMI HeartBeat Missing
   "59_COMMS_HEALTH_DATA"."BRIGE HMI HB ON TIMER".TON(IN := "59_COMMS_HEALTH_DATA"."BRIGE HMI HB", PT := T#1m);
   "59_COMMS_HEALTH_DATA"."BRIGE HMI HB OFF TIMER".TON(IN := NOT "59_COMMS_HEALTH_DATA"."BRIGE HMI HB",
                           PT := T#1m);
END_REGION

REGION Network 14: BRIGE HMI HeartBeat Missing
   RUNG wire#powerrail
      Contact( "59_COMMS_HEALTH_DATA"."BRIGE HMI HB ON TIMER".Q )
      wire#w1
      Coil( "59_COMMS_HEALTH_DATA"."BRIGE HMI HB MISSING" )
   END_RUNG
   RUNG wire#powerrail
      Contact( "59_COMMS_HEALTH_DATA"."BRIGE HMI HB OFF TIMER".Q )
   END_RUNG wire#w1
   // the same network as SCL:
   "59_COMMS_HEALTH_DATA"."BRIGE HMI HB MISSING" := "59_COMMS_HEALTH_DATA"."BRIGE HMI HB ON TIMER".Q OR "59_COMMS_HEALTH_DATA"."BRIGE HMI HB OFF TIMER".Q;
END_REGION
END_FUNCTION

// folder: 500 - 699 Standard FBs

FUNCTION_BLOCK "500_SEQ_STEP"   // FB500, LAD
{ S7_Optimized_Access := 'TRUE' }
VERSION : 0.1
   VAR_INPUT
      SN : Int;   // Step number
      CS : Int;   // Current step
      MST : Time;   // Maximum step time
      SC : Bool;   // Step complete
      BPFLT : Bool;   // Bypass fault
   END_VAR
   VAR_OUTPUT
      ACT : Bool;   // Active
      DN : Bool;   // Done
   END_VAR
   VAR_IN_OUT
      AMST : Time;   // Actual maximum step time
      FLT : Bool;   // Timed out
   END_VAR
   VAR
      RNG : Bool;   // Running
   END_VAR
   VAR RETAIN
      STP_MAX_TIM : TON_TIME;   // Maximum step time
   END_VAR
   VAR
      IEC_Timer_0_Instance : TOF_TIME;
   END_VAR
BEGIN

REGION Network 1: Step Active
   // When step number is active, it is also running
